FUNCTION_BLOCK "CPG_ParetoAnalysis"   // FB31610, SCL
TITLE = CPG_ParetoAnalysis
{ S7_Optimized_Access := 'TRUE' }
AUTHOR : tech.team.motioncontrol@siemens.com
FAMILY : CPG
VERSION : 1.1
// Support: tech.team.motioncontrol@siemens.com
   VAR_INPUT
      ID : DInt;   // ID of the current alarm (0 if no alarm active)
      message : String[40];   // Text of the current alarm
      resetPareto : Bool;   // Rising edge resets statistics
      sort : Int;   // Choose metric to sort by (0=totalDowntime, 1=percentOccurred, 2=timesOccurred, 3=MTTR)
   END_VAR
   VAR_OUTPUT
      totalStops : UInt;   // Total stops due to all faults
      totalTimeSinceReset : Real;   // Total time in minutes since reset
      totalUptime : Real;   // Total uptime in minutes
      totalDowntime : Real;   // Total downtime in minutes
      percentUptime : Real;   // Percent of total time since reset that was uptime
      MTTR : Real;   // Mean time to return
      MTBF : Real;   // Mean time between failures
   END_VAR
   VAR_IN_OUT
      paretoData : Array[0.."CPG_PARTEO_NO_OF_ERRORS_UPPER_LIM"] of "CPG_typePareto";   // Alarm data structure
   END_VAR
   VAR
      statFirstScan : Bool := TRUE;   // Indicate first scan
      statStopReasonOld : DInt;   // The last stop reason
      statResetParetoOld : Bool;   // Reset on the rising edge of resetPareto
      statEntryFound : Bool;   // Alarm code exists already
      statCurrentTimestamp : DTL;   // Current local time
      statPrevTimestamp : DTL;   // Previous local time stamp
      statResetTimestamp : DTL;   // Time when reset
      statSameCurrentTimestamp : Date_And_Time;   // New current time when same alarm is present
      statBaseDowntime : Real;   // Set time when alarm doesn't change
      statIndex : Int;   // Current index in the alarm array
      statTotalStops : UInt;   // Total number of alarm stops
      statTotalDowntime : Real;   // Total machine downtime
      statOverallMTTR : Real;   // Overall total downtime/ Total stops
      statPrevTotalUptime : Real;   // Previous total uptime
      instShellSortPareto : "CPG_ShellSortPareto";   // Sort alarm array
      statSort : String[30];   // Sort alarm data
      statPrevSort : Int;   // Sort on the last scan
      instProgramAlarm : Program_Alarm;   // Record alarm
      statAlarm : Bool;   // Alarm is active
      statArrayFull : Bool;   // Array is larger than MAX_AMOUNT_OF_ERRORS
      statFullRunningDowntime : Real;   // Running downtime when array is full
      statFullPrevDowntime : Real;   // Total downtime for all alarms not recorded in the array
   END_VAR
   VAR_TEMP
      tempTimestamp : DTL;
      tempTimeErr : Int;
      tempEntryFound : Bool;
   END_VAR
   VAR CONSTANT
      MS_TO_MIN : Real := 60000.0;   // Convert from milliseconds to minutes
   END_VAR
BEGIN
   //============================================================================================================
   // SIEMENS NV - APC Belgium
   // (c)Copyright 2018 All Rights Reserved
   //------------------------------------------------------------------------------------------------------------
   // Tested with: S7
   // -1500 with FW version V2.5, V2.6
   // Engineering: TIA Portal V15, V15.1
   // Restrictions: ---
   // Requirements: S7-1x00
   // Functionality: Pareto analysis on stop reasons
   //------------------------------------------------------------------------------------------------------------
   // Change log table:
   // Version       Date               Expert in charge        Changes applied
   // 01.00.00      14.10.2018         J.Pieters               Initial Release 
   // 02.00.00      09.05.2019         K.Bartuska              Included text, total downtime, and MTBF
   // 03.00.00      13.09.2019         K.Bartuska, M.Earnest   Included MTTR, custom sort, and continuous downtime updates         
   //============================================================================================================
   // Function : paretoAnalysis
   //============================================================================================================


   //REGION RESET_PARETO_RESULTS
   IF #statFirstScan OR (#resetPareto AND NOT #statResetParetoOld)
   THEN
       FOR #statIndex := 1 TO "CPG_PARTEO_NO_OF_ERRORS_UPPER_LIM" DO
           #paretoData[#statIndex].alarmID := 0;
           #paretoData[#statIndex].percentageOccurred := 0.0;
           #paretoData[#statIndex].timesOccurred := 0;
           #paretoData[#statIndex].alarmMessage := '';
           #paretoData[#statIndex].MTTR := 0.0;
           #paretoData[#statIndex].totalDowntime := 0.0;
       END_FOR;

       #tempTimeErr := RD_LOC_T(#statResetTimestamp);
       #statTotalStops := 0;
       #statTotalDowntime := 0.0;
       #statOverallMTTR := 0.0;
       #statFirstScan := FALSE;
       #statPrevTotalUptime := 0.0;
       #statStopReasonOld := 0;
       #statArrayFull := 0;
       #statFullPrevDowntime := 0.0;

   END_IF;
   // one shot bit
   #statResetParetoOld := #resetPareto;
   //END_REGION

   FOR #statIndex := 1 TO "CPG_PARTEO_NO_OF_ERRORS_UPPER_LIM" DO
       IF #paretoData[#statIndex].alarmID = #ID
       THEN
           #tempEntryFound := TRUE;
       END_IF;
   END_FOR;

   //REGION UPDATE_DOWNTIME  
   //adjust downtime & MTTR

   //For a different alarm
   IF #ID <> #statStopReasonOld
   THEN
       #statPrevTimestamp := #statCurrentTimestamp;
       #tempTimeErr := RD_LOC_T(#statCurrentTimestamp);
       #statBaseDowntime := 0.0;
       #statAlarm := 0;
       #statFullPrevDowntime := #statFullPrevDowntime + #statFullRunningDowntime;
       #statFullRunningDowntime := 0.0;


       //Update downtime when fault is active    
   ELSIF #ID = #statStopReasonOld AND #ID <> 0
   THEN
       #tempTimeErr := RD_LOC_T(#statSameCurrentTimestamp);
       #statAlarm := 1;
       IF #tempEntryFound
       THEN
           FOR #statIndex := 1 TO "CPG_PARTEO_NO_OF_ERRORS_UPPER_LIM" DO
               IF #paretoData[#statIndex].alarmID = #ID
               THEN
                   #paretoData[#statIndex].totalDowntime := #statBaseDowntime + (DINT_TO_REAL(TIME_TO_DINT(T_DIFF(IN1 := #statSameCurrentTimestamp, IN2 := #statCurrentTimestamp))) / #MS_TO_MIN);
                   IF #paretoData[#statIndex].timesOccurred <> 0
                   THEN
                       #paretoData[#statIndex].MTTR := (#paretoData[#statIndex].totalDowntime) / #paretoData[#statIndex].timesOccurred;
                   END_IF;
                   EXIT;
               END_IF;
           END_FOR;
       ELSIF NOT #tempEntryFound AND #statArrayFull
       THEN
           #statFullRunningDowntime := DINT_TO_REAL(TIME_TO_DINT(T_DIFF(IN1 := #statSameCurrentTimestamp, IN2 := #statCurrentTimestamp))) / #MS_TO_MIN;
       END_IF;
   END_IF;
   //END_REGION


   //REGION CREATE_PROGRAM_ALARM
   //create an alarm
   #instProgramAlarm(SIG := #statAlarm,
                  SD_1 := #ID,
                  SD_2 := #message);
   //END_REGION

   //REGION PARETO_MAIN
   // check if an error is active
   IF #ID <> #statStopReasonOld AND (#ID <> 0)
   THEN
       //REGION INCREMENT_EXISTING_ALARM_ID
       IF #tempEntryFound
       THEN
           FOR #statIndex := 1 TO "CPG_PARTEO_NO_OF_ERRORS_UPPER_LIM" DO
               // find if alarm is already defined in list
               IF #paretoData[#statIndex].alarmID = #ID
               THEN
                   #paretoData[#statIndex].timesOccurred := #paretoData[#statIndex].timesOccurred + UINT#1;
                   EXIT; // exit this loop
               END_IF;
           END_FOR;
       ELSIF NOT #tempEntryFound AND #statArrayFull
       THEN
           #statTotalStops := #statTotalStops + 1;
       END_IF;
       //END_REGION

       //REGION ADD_NEW_ALARM_ID
       //If alarm is not defined in list then make a new entry
       IF (NOT #tempEntryFound) AND (NOT #statArrayFull)
       THEN
           FOR #statIndex := 1 TO "CPG_PARTEO_NO_OF_ERRORS_UPPER_LIM" DO

               IF #paretoData[#statIndex].alarmID = 0
               THEN
                   #paretoData[#statIndex].alarmID := #ID;
                   #paretoData[#statIndex].timesOccurred := 1;
                   #paretoData[#statIndex].alarmMessage := #message;
                   #tempEntryFound := TRUE;
                   //Array is now full
                   IF #statIndex = "CPG_PARTEO_NO_OF_ERRORS_UPPER_LIM"
                   THEN
                       #statArrayFull := 1;
                   END_IF;
                   EXIT; // exit this loop
               END_IF;
           END_FOR;
       END_IF;
       //END_REGION
   END_IF;

   IF #ID <> #statStopReasonOld AND #tempEntryFound
   THEN
       //REGION FIND_TOTAL_OCCURED_ALARMS
       // count total number stop has occured
       //initialize alarm counters
       #statTotalStops := 0;
       #statTotalDowntime := 0.0;
       #statOverallMTTR := 0.0;

       FOR #statIndex := 1 TO "CPG_PARTEO_NO_OF_ERRORS_UPPER_LIM" DO
           IF #paretoData[#statIndex].alarmID = #ID
           THEN
               #statBaseDowntime := #paretoData[#statIndex].totalDowntime;
           END_IF;
           IF #paretoData[#statIndex].alarmID <> 0
           THEN
               #statTotalStops := #statTotalStops + #paretoData[#statIndex].timesOccurred;
               #statTotalDowntime := #statTotalDowntime + #paretoData[#statIndex].totalDowntime;
           END_IF;
       END_FOR;

       IF #statTotalStops <> 0
       THEN
           #statOverallMTTR := (#statTotalDowntime + #statFullPrevDowntime + #statFullRunningDowntime) / #statTotalStops;
       END_IF;
       //END_REGION

       //REGION CALCULATE_PRECENTAGE_FOR_EACH_ALARM
       // calculate percentage each alarm occured
       FOR #statIndex := 1 TO "CPG_PARTEO_NO_OF_ERRORS_UPPER_LIM" DO
           IF #paretoData[#statIndex].alarmID <> 0
           THEN
               // avoid division by zero 
               #paretoData[#statIndex].percentageOccurred := SEL(G := #statTotalStops <> 0,
                                                                 IN0 := 0.0,
                                                                 IN1 := ((#paretoData[#statIndex].totalDowntime) / (#statTotalDowntime + #statFullPrevDowntime + #statFullRunningDowntime)) * 100.0);
           END_IF;
       END_FOR;
       //END_REGION
   END_IF;

   //Update downtime and MTTR when fault is still active
   IF #ID = #statStopReasonOld AND #ID <> 0
   THEN
       //REGION FIND_TOTAL_OCCURED_ALARMS
       IF #tempEntryFound
       THEN
           #statTotalDowntime := 0.0;
           FOR #statIndex := 1 TO "CPG_PARTEO_NO_OF_ERRORS_UPPER_LIM" DO
               #statTotalDowntime := #statTotalDowntime + #paretoData[#statIndex].totalDowntime;
           END_FOR;
       END_IF;

       IF #statTotalStops <> 0 THEN
           #statOverallMTTR := (#statTotalDowntime + #statFullPrevDowntime + #statFullRunningDowntime) / #statTotalStops;
       END_IF;

       //END_REGION

       //REGION CALCULATE_PRECENTAGE_FOR_EACH_ALARM
       // calculate percentage each alarm occured
       IF #tempEntryFound
       THEN
           FOR #statIndex := 1 TO "CPG_PARTEO_NO_OF_ERRORS_UPPER_LIM" DO
               IF #paretoData[#statIndex].alarmID <> 0
               THEN
                   // avoid division by zero 
                   #paretoData[#statIndex].percentageOccurred := SEL(G := #statTotalStops <> 0,
                                                                     IN0 := 0.0,
                                                                     IN1 := ((#paretoData[#statIndex].totalDowntime) / (#statTotalDowntime + #statFullPrevDowntime + #statFullRunningDowntime)) * 100.0);
               END_IF;
           END_FOR;
       END_IF;
       //END_REGION
   END_IF;

   //Sort the alarm array
   //REGION SORT_ARRAY_CRITERIA
   IF #sort = 0 THEN
       #statSort := 'totalDowntime';
   ELSIF #sort = 1 THEN
       #statSort := 'percentageOccurred';
   ELSIF #sort = 2 THEN
       #statSort := 'timesOccurred';
   ELSIF #sort = 3 THEN
       #statSort := 'MTTR';
   END_IF;

   // Sort list: most [statSort] alarms on top (index 1)
   IF #statPrevSort <> #sort OR #ID <> #statStopReasonOld
   THEN
       #instShellSortPareto(mode := TRUE,
                           sortBy := #statSort,
                           variantArray := #paretoData);
   END_IF;
   #statPrevSort := #sort;
   //END_REGION

   #statStopReasonOld := #ID;
   //END_REGION

   //REGION SET_OUTPUTS
   //set other outputs
   #totalStops := #statTotalStops;
   #totalDowntime := #statTotalDowntime + #statFullPrevDowntime + #statFullRunningDowntime;
   #MTTR := #statOverallMTTR;

   //compute total shift time, the amount and percent the machine was up
   #tempTimeErr := RD_LOC_T(#tempTimestamp);
   #totalTimeSinceReset := DINT_TO_REAL(TIME_TO_DINT(T_DIFF(IN1 := #tempTimestamp, IN2 := #statResetTimestamp))) / #MS_TO_MIN;

   #totalUptime := 0.0;

   //if a fault is active the uptime should stay at its previous value
   IF #ID = 0 THEN
       #totalUptime := #totalTimeSinceReset - (#statTotalDowntime + #statFullPrevDowntime + #statFullRunningDowntime);
       #statPrevTotalUptime := #totalUptime;
   ELSE
       #totalUptime := #statPrevTotalUptime;
   END_IF;

   //avoid dividing by zero
   IF #statTotalStops = 0 THEN
       #MTBF := #totalUptime;
   ELSE
       #MTBF := #totalUptime / #statTotalStops;
   END_IF;

   #percentUptime := 100.0 * (#totalUptime) / (#totalTimeSinceReset);
   //END_REGION


   //  -------------- END OF LOGIC -------------------------
   ENO := TRUE;   // Set the ENO output
END_FUNCTION_BLOCK

FUNCTION_BLOCK "CPG_ShellSortPareto"   // FB31611, SCL
TITLE = CPG_ShellSortPareto
{ S7_Optimized_Access := 'TRUE' }
AUTHOR : tech.team.motioncontrol@siemens.com
FAMILY : CPG
VERSION : 1.1
// Support: tech.team.motioncontrol@siemens.com
   VAR_INPUT
      mode : Bool;   // True = sort decending, false = sort ascending
      sortBy : String[30];   // Sorting method
   END_VAR
   VAR_OUTPUT
      done : Bool;   // Sort completed
      error : Bool;   // Error while sorting
      statusID : UInt;   // Indicates block in which error occurred
      status : Word;   // Status word
   END_VAR
   VAR_IN_OUT
      variantArray : Variant;   // Array to be sorted
   END_VAR
   VAR
      statOptions : Struct   // Options for sorting alarm array
         totalDowntime : String[30] := 'totalDowntime';
         timesOccurred : String[30] := 'timesOccurred';
         MTTR : String[30] := 'MTTR';
         percentageOccurred : String[30] := 'percentageOccurred';
      END_STRUCT;
   END_VAR
   VAR_TEMP
      tempArrayPareto : Array[1.."CPG_PARTEO_NO_OF_ERRORS_UPPER_LIM"] of "CPG_typePareto";
      tempElementCount : Int;
      tempElementCopyCount : UDInt;
      tempMoveBlkError : Int;
      tempIncrement : Int;
      tempForCounter : Int;
      tempExchangeIndex : Int;
      tempExchangeVariable : "CPG_typePareto";
      tempTypeTag : "CPG_typePareto";
   END_VAR
   VAR CONSTANT
      MAX_ARRAY_ELEMENTS : Int := 1000;
      NO_ERROR : Word := 16#0000;
      NO_CURRENT_JOBS : Word := 16#7000;
      EMPTY_ARRAY : Word := 16#8200;
      NOT_AN_ARRAY : Word := 16#8201;
      WRONG_ELEMENT_TYPE : Word := 16#8202;
      TOO_MANY_ELEMENTS : Word := 16#8203;
      ERROR_IN_THIS_BLOCK : UInt := 1;
      ERROR_MOVE_BLK_VARIANT_R : UInt := 2;
      ERROR_MOVE_BLK_VARIANT_W : UInt := 3;
   END_VAR
BEGIN
   //=============================================================================
   // SIEMENS AG
   // (c)Copyright 2017
   //-----------------------------------------------------------------------------
   // Library:       LGF (Library General Functions)
   // Tested with:   CPU1212C DC/DC/DC FW:V4.2
   // Engineering:   TIA Portal V14 Update 1
   // Restrictions:  -
   // Requirements:  PLC (S7-1200 / S7-1500)
   // Functionality: A shellsort algorithm with a complexity between 'n^2' and
   //                'n log n' for average, best and worst case inputs and space
   //                complexity '1'.
   //                The block accepts a pareto array as an inOut-variable and
   //                returns the sorted version of the array in the same variable
   //-----------------------------------------------------------------------------
   // Change log table:
   // Version  Date        Expert in charge / Changes applied
   // 01.00.00 19.08.2015  Siemens Industry Online Support
   //                      First released version
   // 01.01.00 19.05.2016  Siemens Industry Online Support
   //                      New function: reverse sort
   // 01.01.01 02.01.2017  Siemens Industry Online Support
   //                      Upgrade: TIA Portal V14 Update 1
   // 01.01.02 17.08.2018  Siemens Industry Online Support
   //                      Upgrade: TIA V15 Update 2
   // 01.01.03 26.10.2018  APC-BE - Pieters
   //                      Modified for use with pareto type
   // 01.01.03 13.09.2019  Modified with variable sort parameters                  
   //-----------------------------------------------------------------------------
   //Status Codes:
   // 16#7000:  No current jobs
   // 16#0000:  Job finished; Note: There is no "Busy"-Status because the block is
   //           finished within a single cycle
   // 16#8200:  Error: Parameter is an array with only one element
   // 16#8201:  Error: Parameter is not an array
   // 16#8202:  Error: Parameter is an array of the wrong type
   //           (correct type is Real)
   // 16#8203:  Error: There are too many Elements in the array
   //           (default: max. 1000 Elements)
   //=============================================================================

   // Change note: If you wish to use this shellsort block for other datatypes,
   // you simply need to change the following variables to that type
   // 1. tempExchangeVariable
   // 2. tempTypeTag
   // 3. tempArray<Type>
   // Space note: If you wish to reduce the space of this block, you may reduce the
   // size of the tempArray<Type> to one just big enough for your specific purpose
   // It is not recommended to increase the size significantly.

   // Initialization
   #tempElementCount := 0;
   #tempElementCopyCount := 0;
   #tempMoveBlkError := 0;
   #tempIncrement := 0;
   #tempForCounter := 0;
   #tempExchangeIndex := 0;
   #tempExchangeVariable.alarmID := 0;
   #tempExchangeVariable.percentageOccurred := 0.0;
   #tempExchangeVariable.timesOccurred := 0;
   #tempTypeTag.alarmID := 0;
   #tempTypeTag.percentageOccurred := 0.0;
   #tempTypeTag.timesOccurred := 0;

   // Set "No current job" status
   #done := false;
   #error := false;
   #statusID := #ERROR_IN_THIS_BLOCK;
   #status := #NO_CURRENT_JOBS;


   // If the variant inOut-parameter is not an array, set error status 8201
   IF (IS_ARRAY(#variantArray) = false) THEN
       #error := true;
       #statusID := #ERROR_IN_THIS_BLOCK;
       #status := #NOT_AN_ARRAY;
       RETURN;
   ELSE
       IF TypeOfElements(#variantArray) = TypeOf(#tempTypeTag) THEN
           // If the parameter is an array of the type real, get the element count
           #tempElementCopyCount := CountOfElements(#variantArray);
           #tempElementCount := UDINT_TO_INT(CountOfElements(#variantArray));
           // Check whether the variant array contains less than the maximum possible amount of elements
           IF #tempElementCount > #MAX_ARRAY_ELEMENTS THEN
               #error := true;
               #statusID := #ERROR_IN_THIS_BLOCK;
               #status := #TOO_MANY_ELEMENTS;
               RETURN;
           END_IF;
       ELSE
           // If the parameter is an array but not of the type real, set an error status
           #error := true;
           #statusID := #ERROR_IN_THIS_BLOCK;
           #status := #WRONG_ELEMENT_TYPE;
           RETURN;
       END_IF;
   END_IF;

   // If there are more than zero elements to sort, begin sorting    
   IF #tempElementCount > 1 AND #error = false THEN

       // Read the elements of the incoming variant-array and write into the local array
       #tempMoveBlkError := MOVE_BLK_VARIANT(COUNT := #tempElementCopyCount,
                                             DEST => #tempArrayPareto,
                                             DEST_INDEX := 0,
                                             SRC := #variantArray,
                                             SRC_INDEX := 0);

       // Error handling for MOVE_BLK_VARIANT
       IF #tempMoveBlkError <> 0 THEN
           #error := true;
           #statusID := #ERROR_MOVE_BLK_VARIANT_R;
           #status := INT_TO_WORD(#tempMoveBlkError);
           RETURN;
       END_IF;

       // ShellSort Start
       #tempIncrement := 1;
       REPEAT
           #tempIncrement := (3 * #tempIncrement) + 1;
       UNTIL #tempIncrement > #tempElementCount
       END_REPEAT;

       REPEAT
           #tempIncrement := DINT_TO_INT(TRUNC(#tempIncrement / 3));
           FOR #tempForCounter := (#tempIncrement + 1) TO #tempElementCount DO
               #tempExchangeVariable := #tempArrayPareto[#tempForCounter];
               #tempExchangeIndex := #tempForCounter;

               IF #mode  // Modification Version 02.00.00
               THEN      //mode = TRUE --> sort descending  
                   //Downtime
                   IF #sortBy = #statOptions.totalDowntime THEN
                       WHILE ((#tempArrayPareto[#tempExchangeIndex - #tempIncrement].totalDowntime < #tempExchangeVariable.totalDowntime)) DO
                           #tempArrayPareto[#tempExchangeIndex] := #tempArrayPareto[#tempExchangeIndex - #tempIncrement];
                           #tempExchangeIndex := #tempExchangeIndex - #tempIncrement;
                           IF (#tempExchangeIndex <= #tempIncrement) THEN
                               GOTO EXITWhile;
                           END_IF;
                       END_WHILE;
                       //Times Occurred    
                   ELSIF #sortBy = #statOptions.timesOccurred THEN
                       WHILE ((#tempArrayPareto[#tempExchangeIndex - #tempIncrement].timesOccurred < #tempExchangeVariable.timesOccurred)) DO
                           #tempArrayPareto[#tempExchangeIndex] := #tempArrayPareto[#tempExchangeIndex - #tempIncrement];
                           #tempExchangeIndex := #tempExchangeIndex - #tempIncrement;
                           IF (#tempExchangeIndex <= #tempIncrement) THEN
                               GOTO EXITWhile;
                           END_IF;
                       END_WHILE;
                       //Percentage Occurred
                   ELSIF #sortBy = #statOptions.percentageOccurred THEN
                       WHILE ((#tempArrayPareto[#tempExchangeIndex - #tempIncrement].percentageOccurred < #tempExchangeVariable.percentageOccurred)) DO
                           #tempArrayPareto[#tempExchangeIndex] := #tempArrayPareto[#tempExchangeIndex - #tempIncrement];
                           #tempExchangeIndex := #tempExchangeIndex - #tempIncrement;
                           IF (#tempExchangeIndex <= #tempIncrement) THEN
                               GOTO EXITWhile;
                           END_IF;
                       END_WHILE;
                       // MTTR
                   ELSIF #sortBy = #statOptions.MTTR THEN
                       WHILE ((#tempArrayPareto[#tempExchangeIndex - #tempIncrement].MTTR < #tempExchangeVariable.MTTR)) DO
                           #tempArrayPareto[#tempExchangeIndex] := #tempArrayPareto[#tempExchangeIndex - #tempIncrement];
                           #tempExchangeIndex := #tempExchangeIndex - #tempIncrement;
                           IF (#tempExchangeIndex <= #tempIncrement) THEN
                               GOTO EXITWhile;
                           END_IF;
                       END_WHILE;
                   END_IF;

               ELSE      // mode = FALSE --> sort ascending
                   WHILE ((#tempArrayPareto[#tempExchangeIndex - #tempIncrement].MTTR > #tempExchangeVariable.MTTR)) DO
                       #tempArrayPareto[#tempExchangeIndex] := #tempArrayPareto[#tempExchangeIndex - #tempIncrement];
                       #tempExchangeIndex := #tempExchangeIndex - #tempIncrement;
                       IF (#tempExchangeIndex <= #tempIncrement) THEN
                           GOTO EXITWhile;
                       END_IF;
                   END_WHILE;
               END_IF;

           EXITWhile:
               #tempArrayPareto[#tempExchangeIndex] := #tempExchangeVariable;
           END_FOR;
       UNTIL #tempIncrement <= 1
       END_REPEAT;
       // ShellSort End

       // Write the elements of the local array back to the variant array
       #tempMoveBlkError := MOVE_BLK_VARIANT(COUNT := #tempElementCopyCount,
                                             DEST => #variantArray,
                                             DEST_INDEX := 0,
                                             SRC := #tempArrayPareto,
                                             SRC_INDEX := 0);

       // Error handling for MOVE_BLK_VARIANT
       IF #tempMoveBlkError <> 0 THEN
           #statusID := #ERROR_MOVE_BLK_VARIANT_W;
           #status := INT_TO_WORD(#tempMoveBlkError);
           RETURN;
       END_IF;

       // Set output status = "Job Finished" and output Done = true
       #done := true;
       #status := #NO_ERROR;

   ELSIF #tempElementCount <= 1 THEN
       // If there are 0 elements in the array, set status to "Error: Parameter is an empty array"
       #error := true;
       #statusID := #ERROR_IN_THIS_BLOCK;
       #status := #EMPTY_ARRAY;
   END_IF;

   //  -------------- END OF LOGIC -------------------------
   ENO := TRUE;   // Set the ENO output
END_FUNCTION_BLOCK

FUNCTION_BLOCK "CPG_RecipeControl"   // FB31612, SCL
TITLE = CPG_RecipeControl
{ S7_Optimized_Access := 'TRUE' }
AUTHOR : tech.team.motioncontrol@siemens.com
FAMILY : CPG
VERSION : 1.1
// Support: tech.team.motioncontrol@siemens.com
   VAR_INPUT
      enable : Bool;   // Recipe change is only possible if instruction is enabled
      recipeChangeID : Int;   // ID of recipe to change to
      recipeChangeReq : Bool;   // Change recipe on rising edge
      recipeSaveReq : Bool;   // Save current recipe on rising edge
      recipeSaveAsID : Int;   // Location to saveas recipe to
      recipeSaveAsReq : Bool;   // SaveAs recipe on rising edge
      recipeCopySourceID : Int;   // Location to copy recipe from
      recipeCopyID : Int;   // Location to copy recipe to
      recipeCopyReq : Bool;   // Copy recipe on rising edge
      newRecipeName : String[60];   // Name of the saveas or copied recipe
      recipeDeleteID : Int;   // Location of recipe to delete
      recipeDeleteReq : Bool;   // Delete recipe on rising edge
      resetAllTimes : Bool;   // Reset cumulative seconds for all recipes
   END_VAR
   VAR_OUTPUT
      currentRecipeID : Int;   // ID of the current recipe
      currentRecipeName : String[60];   // Name of the current recipe
      recipeChangeDisabled : Bool;   // Recipe changes are enabled
      recipeSetpointDiff : Bool;   // New setpoint differs from current recipe value
      recipeCurrentSeconds : Time;   // Current recipe time in seconds
      error : Bool;   // Error Present
      errorID : Word := 16#0000;   // Code for Status
   END_VAR
   VAR_IN_OUT
      recipeControl : "CPG_typeRecipeControl";   // Recipe Control tag
      recipeNames : Array[0.."CPG_NO_OF_RECIPE_UPPER_LIM"] of String[60];   // All recipe names
      recipeCumSeconds : Array[0.."CPG_NO_OF_RECIPE_UPPER_LIM"] of Time;   // Cumulative times for all recipes
      recipeSaveDates : Array[0.."CPG_NO_OF_RECIPE_UPPER_LIM"] of DTL;   // Recipe saved date time
   END_VAR
   VAR
      statSetpoinDiffTimer : TON_TIME;
      statPrevRecipe : Int;
      statChangeReq : R_TRIG;
      statSaveReq : R_TRIG;
      statSaveAsReq : R_TRIG;
      statCopyReq : R_TRIG;
      statDeleteReq : R_TRIG;
      statChangeTimer : TP_TIME;
      statChangeTimerFall : F_TRIG;
      statSaveTimer : TP_TIME;
      statSaveTimerFall : F_TRIG;
      statSaveAsTimer : TP_TIME;
      statSaveAsTimerFall : F_TRIG;
      statCopyTimer : TP_TIME;
      statCopyTimerFall : F_TRIG;
      statDeleteTimer : TP_TIME;
      statDeleteTimerFall : F_TRIG;
      statPrevCumSeconds : Array[0.."CPG_NO_OF_RECIPE_UPPER_LIM"] of Time;
      statChangeTimeStamp : DTL;
   END_VAR
   VAR_TEMP
      tempChangeEN : Bool;
      tempCopyRecipeEN : Bool;
      tempSaveRecipeEN : Bool;
      tempDeleteRecipeEN : Bool;
      tempDTLError : Int;
      tempLoop : Int;
      tempTime : DTL;
      tempRecipeSaveAs : Bool;
   END_VAR
   VAR CONSTANT
      MAX_RECIPE_NUM : Int := 20;
      WARNING_TIMERLEN : Time := T#1s;
      CHG_ERR : Word := 16#8001;
      SAVE_ERR : Word := 16#8002;
      COPY_ERR : Word := 16#8004;
      DEL_ERR : Word := 16#8008;
   END_VAR
BEGIN
   //============================================================================================================
   // SIEMENS AG
   // (c)Copyright 2019 All Rights Reserved
   //------------------------------------------------------------------------------------------------------------
   // Library: LCPG
   // Tested with: S7-1500 with FW version V2.1
   // Engineering: TIA Portal V14
   // Restrictions: ---
   // Requirements: S7-1500
   // Functionality: used to control the current machine recipe
   // Support: tech.team.motioncontrol@siemens.com
   //------------------------------------------------------------------------------------------------------------
   // Change log table:
   // Version       Date               Expert in charge    Changes applied
   //  01.01.00     02.01.2019         KB                  Initial Release
   //============================================================================================================
   // Function : CPG_RecipeControl
   //============================================================================================================

   REGION INITIALIZATION
       #errorID := 16#0000;

       #recipeControl.RecipeChangeDisabled := NOT #enable;

       //check lanugage for out of bounds
       IF (#recipeControl.LanguageSelection < 0) OR (#recipeControl.LanguageSelection > "LPMLV30_LANGUAGES_UPPER_LIM") THEN
           #errorID := #errorID OR 16#1000;
           #recipeControl.LanguageSelection := 0;
       END_IF;


       //Dectect any recipe & setpoint differences
       //if any call of recipe setpoint FBs has a difference, the RecipeSetpointDiff bit is set
       IF #recipeControl.RecipeSetpointDiff THEN
           #recipeSetpointDiff := true;
           #recipeControl.RecipeSetpointDiff := false;
       END_IF;
   END_REGION


   REGION RECIPE MANAGEMENT ENABLING
       //Check that only 1 recipe command is active
       IF NOT (#recipeControl.RecipeCopy OR #recipeControl.RecipeDelete OR #recipeControl.RecipeSave) THEN     //all false except change
           #tempChangeEN := true;
       END_IF;
       IF NOT (#recipeControl.RecipeCopy OR #recipeControl.RecipeDelete OR #recipeControl.RecipeChange) THEN   //all false except save/saveas
           #tempSaveRecipeEN := true;
       END_IF;
       IF NOT (#recipeControl.RecipeChange OR #recipeControl.RecipeDelete OR #recipeControl.RecipeSave) THEN   //all false except copy
           #tempCopyRecipeEN := true;
       END_IF;
       IF NOT (#recipeControl.RecipeCopy OR #recipeControl.RecipeChange OR #recipeControl.RecipeSave) THEN     //all false except delete
           #tempDeleteRecipeEN := true;
       END_IF;


       //RecipeCmd out of bounds, or equal to the current recipe
       IF (#recipeChangeID > #MAX_RECIPE_NUM) OR (#recipeChangeID < 0) OR (#recipeChangeID = #recipeControl.CurrentRecipeID) THEN
           #errorID := #errorID OR #CHG_ERR;
           #tempChangeEN := false;
       END_IF;
       //RecipeSaveAsCmd out of bounds, or attempting to over current recipe
       IF (#recipeSaveAsID > #MAX_RECIPE_NUM) OR (#recipeSaveAsID < 0) OR (#recipeSaveAsID = #recipeControl.CurrentRecipeID) THEN
           #errorID := #errorID OR #SAVE_ERR;
           #tempSaveRecipeEN := false;
       END_IF;
       //RecipeCopyCmd or RecipeCopySourceCmd out of bounds, cannot copy to currently running recipe
       IF (#recipeCopyID > #MAX_RECIPE_NUM) OR (#recipeCopyID < 0) OR (#recipeCopySourceID > #MAX_RECIPE_NUM) OR (#recipeCopySourceID < 0)
           OR #recipeCopyID = #recipeControl.CurrentRecipeID THEN
           #errorID := #errorID OR #COPY_ERR;
           #tempCopyRecipeEN := false;
       END_IF;
       //RecipeDeleteCmd out of bounds or equal to current recipe
       IF (#recipeDeleteID > #MAX_RECIPE_NUM) OR (#recipeDeleteID < 0) OR (#recipeDeleteID = #recipeControl.CurrentRecipeID) THEN
           #errorID := #errorID OR #DEL_ERR;
           #tempDeleteRecipeEN := false;
       END_IF;
   END_REGION


   REGION RECIPE CHANGE
       //only allow recipe changes while enabled
       IF #enable THEN

           //timer needed for display & troubleshooting
           //timer starts on rising edge of the req signal and persists for 1s
           #statChangeReq(CLK := #recipeChangeReq);

           #statChangeTimer(IN := #statChangeReq.Q,
                        PT := #WARNING_TIMERLEN);

           #statChangeTimerFall(CLK := #statChangeTimer.Q);


           //Check that the recipe to change is valid & no other command is active
           IF #tempChangeEN THEN

               //set output to indicate that a recipe is being changed
               IF #statChangeTimer.Q THEN
                   #recipeControl.RecipeChange := true;
               ELSE
                   #recipeControl.RecipeChange := false;
               END_IF;

               //change recipe on done bit, true for only 1 scan
               IF #statChangeTimerFall.Q THEN
                   #recipeControl.RecipeChangeNum := #recipeControl.RecipeChangeNum + 1;
                   #recipeControl.CurrentRecipeID := #recipeChangeID;
                   #recipeControl.CurrentRecipeName := #recipeNames[#recipeControl.CurrentRecipeID];
               END_IF;

           END_IF;

       END_IF;
   END_REGION


   REGION RECIPE SAVEAS
       //timer needed for display & troubleshooting
       //timer starts on rising edge of the req signal and persists for 1s
       #statSaveAsReq(CLK := #recipeSaveAsReq);

       #statSaveAsTimer(IN := #statSaveAsReq.Q,
                    PT := #WARNING_TIMERLEN);

       #statSaveAsTimerFall(CLK := #statSaveAsTimer.Q);


       //Check that the recipe to save is valid & no other command is active
       IF #tempSaveRecipeEN THEN

           //set output to indicate that a recipe is being saved
           //because Save & SaveAs use the same output (RecipeControl.RecipeSave), this is handled slightly differently
           IF #statSaveAsTimer.Q THEN
               #tempRecipeSaveAs := true;
           END_IF;


           //set work variables so that setpoints know the source/destination of the copy operation
           IF #statSaveAsTimer.Q THEN
               #recipeControl.RecipeSourceID := #recipeControl.CurrentRecipeID;
               #recipeControl.RecipeDestinationID := #recipeSaveAsID;
           END_IF;

           //update counter, take timestamp, and update recipe name
           IF #statSaveAsTimerFall.Q THEN
               #recipeControl.RecipeSaveNum := #recipeControl.RecipeSaveNum + 1;
               #tempDTLError := RD_LOC_T(#recipeSaveDates[#recipeControl.RecipeDestinationID]);
               #recipeNames[#recipeControl.RecipeDestinationID] := #newRecipeName;
           END_IF;

       END_IF;
   END_REGION


   REGION RECIPE SAVE
       //timer needed for display & troubleshooting
       //timer starts on rising edge of the req signal and persists for 1s
       #statSaveReq(CLK := #recipeSaveReq);

       #statSaveTimer(IN := #statSaveReq.Q,
                  PT := #WARNING_TIMERLEN);

       #statSaveTimerFall(CLK := #statSaveTimer.Q);


       //saving is always possible
       //note that the saveas REGION must be after the save REGION
       //otherwise RecipeControl.RecipeSave won't be set by a saveas

       //set output to indicate that a recipe is being saved
       //because Save & SaveAs use the same output (RecipeControl.RecipeSave), this is handled slightly differently
       IF #statSaveTimer.Q  OR #tempRecipeSaveAs THEN
           #recipeControl.RecipeSave := true;
       ELSE
           #recipeControl.RecipeSave := false;
       END_IF;

       //set work variables so that setpoints know the source/destination of the save operation
       IF #statSaveTimer.Q THEN
           #recipeControl.RecipeSourceID := #recipeControl.CurrentRecipeID;
           #recipeControl.RecipeDestinationID := #recipeControl.CurrentRecipeID;
       END_IF;

       //update counter, take timestamp
       IF #statSaveTimerFall.Q THEN
           #recipeControl.RecipeSaveNum := #recipeControl.RecipeSaveNum + 1;
           #tempDTLError := RD_LOC_T(#recipeSaveDates[#recipeControl.RecipeDestinationID]);
       END_IF;
   END_REGION


   REGION RECIPE COPY
       //timer needed for display & troubleshooting
       //timer starts on rising edge of the req signal and persists for 1s
       #statCopyReq(CLK := #recipeCopyReq);

       #statCopyTimer(IN := #statCopyReq.Q,
                  PT := #WARNING_TIMERLEN);

       #statCopyTimerFall(CLK := #statCopyTimer.Q);


       //Check that the recipes to copy are valid & no other command is active
       IF #tempCopyRecipeEN THEN

           //set output to indicate that a recipe is being copied
           IF #statCopyTimer.Q THEN
               #recipeControl.RecipeCopy := true;
           ELSE
               #recipeControl.RecipeCopy := false;
           END_IF;

           //set work variables so that setpoints know the source/destination of the copy operation
           IF #statCopyTimer.Q THEN
               #recipeControl.RecipeSourceID := #recipeCopySourceID;
               #recipeControl.RecipeDestinationID := #recipeCopyID;
           END_IF;

           //update the recipename of the new recipe, increment change work variable
           IF #statCopyTimerFall.Q THEN
               #recipeControl.RecipeCopyNum := #recipeControl.RecipeCopyNum + 1;
               #tempDTLError := RD_LOC_T(#recipeSaveDates[#recipeControl.RecipeDestinationID]);
               #recipeNames[#recipeControl.RecipeDestinationID] := #newRecipeName;
           END_IF;

       END_IF;
   END_REGION


   REGION RECIPE DELETE
       //timer needed for display & troubleshooting
       //timer starts on rising edge of the req signal and persists for 1s
       #statDeleteReq(CLK := #recipeDeleteReq);

       #statDeleteTimer(IN := #statDeleteReq.Q,
                    PT := #WARNING_TIMERLEN);

       #statDeleteTimerFall(CLK := #statDeleteTimer.Q);


       //Check that the recipe to delete is valid & no other command is active
       IF #tempDeleteRecipeEN THEN

           //set output to indicate that a recipe is being copied
           IF #statDeleteTimer.Q THEN
               #recipeControl.RecipeDelete := true;
           ELSE
               #recipeControl.RecipeDelete := false;
           END_IF;

           //set work variable so that setpoints know the destination of the delete operation
           IF #statDeleteTimer.Q THEN
               #recipeControl.RecipeDestinationID := #recipeDeleteID;
           END_IF;

           //clear the recipe name
           IF #statDeleteTimerFall.Q THEN
               #recipeControl.RecipeDeleteNum := #recipeControl.RecipeDeleteNum + 1;
               #tempDTLError := RD_LOC_T(#recipeSaveDates[#recipeControl.RecipeDestinationID]);
               #recipeNames[#recipeControl.RecipeDestinationID] := '';
           END_IF;

       END_IF;
   END_REGION


   REGION TIME TRACKING
       //reset all times resets the cumulative time for all recipes, and the cum seconds output, but does not change the save timestamps
       IF #resetAllTimes THEN
           FOR #tempLoop := 0 TO #MAX_RECIPE_NUM DO
               // set all cumulative times to zero
               #recipeCumSeconds[#tempLoop] := T#0s;
               #statPrevCumSeconds[#tempLoop] := T#0s;
           END_FOR;
           #recipeCurrentSeconds := T#0s;
       END_IF;

       //if recipe changes, note the time of change and save the accumulated time for the 
       IF #recipeControl.CurrentRecipeID <> #statPrevRecipe THEN
           #tempDTLError := RD_LOC_T(#statChangeTimeStamp);
           #statPrevCumSeconds[#recipeControl.CurrentRecipeID] := #recipeCumSeconds[#recipeControl.CurrentRecipeID];
           #recipeCurrentSeconds := T#0s;
       END_IF;

       //must initialize this value or timetracking does not work on plc startup
       IF #statChangeTimeStamp = DTL#1970-01-01-00:00:00 THEN
           #tempDTLError := RD_LOC_T(#statChangeTimeStamp);
       END_IF;

       #tempDTLError := RD_LOC_T(#tempTime);
       #recipeCurrentSeconds := T_DIFF(IN1 := #tempTime, IN2 := #statChangeTimeStamp);
       #recipeCumSeconds[#recipeControl.CurrentRecipeID] := #statPrevCumSeconds[#recipeControl.CurrentRecipeID] + #recipeCurrentSeconds;
   END_REGION


   REGION SET OUTPUTS
       //Update current recipe name in case user changed RecipeControl.CurrentRecipeName on the HMI
       IF #recipeControl.CurrentRecipeName <> #recipeNames[#recipeControl.CurrentRecipeID] THEN
           #recipeNames[#recipeControl.CurrentRecipeID] := #recipeControl.CurrentRecipeName;
       ELSE
           #recipeControl.CurrentRecipeName := #recipeNames[#recipeControl.CurrentRecipeID];
       END_IF;

       //tmpDTLerror recieves a value if there is an eror returning the PLC system time
       IF #tempDTLError <> 0 THEN
           #errorID := #errorID OR 16#0100;
       END_IF;

       //report error bit
       IF #errorID = 16#0 THEN
           #error := false;
       ELSE
           #error := true;
       END_IF;

       //ensure recipe display numbers are in bounds
       #recipeControl.RecipeID_A := LIMIT(MN := 0, IN := #recipeControl.RecipeID_A, MX := #MAX_RECIPE_NUM);
       #recipeControl.RecipeID_B := LIMIT(MN := 0, IN := #recipeControl.RecipeID_B, MX := #MAX_RECIPE_NUM);
       #recipeControl.RecipeID_C := LIMIT(MN := 0, IN := #recipeControl.RecipeID_C, MX := #MAX_RECIPE_NUM);

       //set some final outputs
       #statPrevRecipe := #recipeControl.CurrentRecipeID;
       #currentRecipeID := #recipeControl.CurrentRecipeID;
       #currentRecipeName := #recipeControl.CurrentRecipeName;
       #recipeChangeDisabled := #recipeControl.RecipeChangeDisabled;
   END_REGION

   //  -------------- END OF LOGIC -------------------------
   ENO := TRUE;   // Set the ENO output
END_FUNCTION_BLOCK

FUNCTION_BLOCK "CPG_RecipeHMIManager"   // FB31613, SCL
TITLE = CPG_RecipeHMIManager
{ S7_Optimized_Access := 'TRUE' }
AUTHOR : tech.team.motioncontrol@siemens.com
FAMILY : CPG
VERSION : 1.1
// Support: tech.team.motioncontrol@siemens.com
   VAR_INPUT
      recipePopupTrackers : Array[0..#NUM_TYPES] of Int;   // Index of recipe that is to be displayed in popup
   END_VAR
   VAR_OUTPUT
      setpointsArray_REAL : Array[0..11] of "CPG_typeRecipeSetpoint_REAL";   // Setpoints to display
      setpointsArray_DINT : Array[0..11] of "CPG_typeRecipeSetpoint_DINT";   // Setpoints to display
      setpointsArray_BOOL : Array[0..11] of "CPG_typeRecipeSetpoint_BOOL";   // Setpoints to display
      setpointsArray_STRING : Array[0..11] of "CPG_typeRecipeSetpoint_STRING";   // Setpoints to display
      recipeMaxPages : Array[0..4] of Int;   // Max pages for all types of setpoint
      setpointFaceplatesDisable_REAL : Array[0..11] of Bool;   // True if that setpoint should be hidden
      "setpoint FaceplatesDisable_DINT" : Array[0..11] of Bool;   // True if that setpoint should be hidden
      "setpoint FaceplatesDisable_BOOL" : Array[0..11] of Bool;   // True if that setpoint should be hidden
      "setpoint FaceplatesDisable_STRING" : Array[0..11] of Bool;   // True if that setpoint should be hidden
      recipeArrayNames : Array[0..19] of String[60];   // Recipe names to display
      recipeArraySaves : Array[0..19] of DTL;   // Recipe save times to display
      recipeArrayTimes : Array[0..19] of Time;   // Recipe cumtimes to display
      recipeArrayDisables : Array[0..19] of Bool;   // True if that recipe should be hidden
      recipeArrayNums : Array[0..19] of Int;   // Recipe numbers to display
   END_VAR
   VAR_IN_OUT
      setpoints_REAL : Array[*] of "CPG_typeRecipeSetpoint_REAL";   // Machine setpoints
      setpoints_DINT : Array[*] of "CPG_typeRecipeSetpoint_DINT";   // Machine setpoints
      setpoints_BOOL : Array[*] of "CPG_typeRecipeSetpoint_BOOL";   // Machine setpoints
      setpoints_STRING : Array[*] of "CPG_typeRecipeSetpoint_STRING";   // Machine setpoints
      recipePopup_REAL : "CPG_typeRecipeSetpoint_REAL";   // Tag of popup
      recipePopup_DINT : "CPG_typeRecipeSetpoint_DINT";   // Tag of popup
      recipePopup_BOOL : "CPG_typeRecipeSetpoint_BOOL";   // Tag of popup
      recipePopup_STRING : "CPG_typeRecipeSetpoint_STRING";   // Tag of popup
      recipeCurrentPages : Array[0..4] of Int;   // Current page for viewing setpoints/recipies
      recipeNamesArray : Array[*] of String[60];   // Recipe names
      recipeSavesArray : Array[*] of DTL;   // Recipe saves
      recipeTimesArray : Array[*] of Time;   // Recipe cumtimes
   END_VAR
   VAR
      statPrevCurrentPages : Array[0..4] of Int;
      statPrevPopupTrackers : Array[0..#NUM_TYPES] of Int;
      statPrevPopupsSave : Array[0..#NUM_TYPES] of Bool;
      statPrevPopupsRevert : Array[0..#NUM_TYPES] of Bool;
      statPrevPopupIN_REAL : Real;
      statPrevSetpointIN_REAL : Real;
      statPrevPopupIN_DINT : DInt;
      statPrevSetpointIN_DINT : DInt;
      statPrevPopupIn_BOOL : Bool;
      statPrevSetpointIn_BOOL : Bool;
      statPrevPopupIn_STRING : String[60];
      statPrevSetpointIn_STRING : String[60];
   END_VAR
   VAR_TEMP
      tempLoop : Int;
      tempSetptsLower : Array[0..#NUM_TYPES] of Int;
      tempSetptsUpper : Array[0..#NUM_TYPES] of Int;
      tempCurrentPopup : Int;
      tempNumRecipesLower : Int;
      tempNumRecipesUpper : Int;
   END_VAR
   VAR CONSTANT
      NUM_TYPES : Int := 3;
      SETPOINTS_PERPAGE : Int := 12;
      RECIPES_PERPAGE : Int := 20;
      INDEX_REAL : Int := 0;
      INDEX_DINT : Int := 1;
      INDEX_BOOL : Int := 2;
      INDEX_STRING : Int := 3;
   END_VAR
   // statPrevCurrentPages[0] := -1;
   // statPrevCurrentPages[1] := -1;
   // statPrevCurrentPages[2] := -1;
   // statPrevCurrentPages[3] := -1;
   // statPrevPopupTrackers[0] := -1;
   // statPrevPopupTrackers[1] := -1;
   // statPrevPopupTrackers[2] := -1;
   // statPrevPopupTrackers[3] := -1;
BEGIN
   //============================================================================================================
   // SIEMENS AG
   // (c)Copyright 2019 All Rights Reserved
   //------------------------------------------------------------------------------------------------------------
   // Library: LCPG
   // Tested with: S7-1500 with FW version V2.1
   // Engineering: TIA Portal V14
   // Restrictions: ---
   // Requirements: S7-1500
   // Functionality: handles the automatic display of setpoints/recipies
   // Support: tech.team.motioncontrol@siemens.com
   //------------------------------------------------------------------------------------------------------------
   // Change log table:
   // Version       Date               Expert in charge    Changes applied
   //  01.01.00     02.01.2019         KB                  Initial Release
   //============================================================================================================
   // Function : CPG_RecipeHMIManager
   //============================================================================================================
   //

   //This function handles the automatic display of the four types of setpoints and the list of recipies
   //There can be any number of setpoints or recipies, but only 12 setpoints and 20 recipies will fit on the screen
   //This block copies 12 of the setpoints into an auxillary array, which is actually displayed on the screen
   //Which 12 setpoints are copied depends on the current page
   //A similar procedure is carried out for the 20 recipe names displayed on the "Recipe_Control" screen
   //Lastly, the recipe that's currently selected is loaded into the popup tag,
   //and any changes made to that tag are propogated back into the "true" setpoint tag
   //The user generally will not need to modify the contents of this block


   REGION CALCULATE BOUNDS
       //calculate upper and lower limits 
       #tempSetptsLower[0] := DINT_TO_INT(LOWER_BOUND(ARR := #setpoints_REAL, DIM := 1));
       #tempSetptsLower[1] := DINT_TO_INT(LOWER_BOUND(ARR := #setpoints_DINT, DIM := 1));
       #tempSetptsLower[2] := DINT_TO_INT(LOWER_BOUND(ARR := #setpoints_BOOL, DIM := 1));
       #tempSetptsLower[3] := DINT_TO_INT(LOWER_BOUND(ARR := #setpoints_STRING, DIM := 1));
       #tempNumRecipesLower := DINT_TO_INT(LOWER_BOUND(ARR := #recipeNamesArray, DIM := 1));

       #tempSetptsUpper[0] := DINT_TO_INT(UPPER_BOUND(ARR := #setpoints_REAL, DIM := 1));
       #tempSetptsUpper[1] := DINT_TO_INT(UPPER_BOUND(ARR := #setpoints_DINT, DIM := 1));
       #tempSetptsUpper[2] := DINT_TO_INT(UPPER_BOUND(ARR := #setpoints_BOOL, DIM := 1));
       #tempSetptsUpper[3] := DINT_TO_INT(UPPER_BOUND(ARR := #setpoints_STRING, DIM := 1));
       #tempNumRecipesUpper := DINT_TO_INT(UPPER_BOUND(ARR := #recipeNamesArray, DIM := 1));